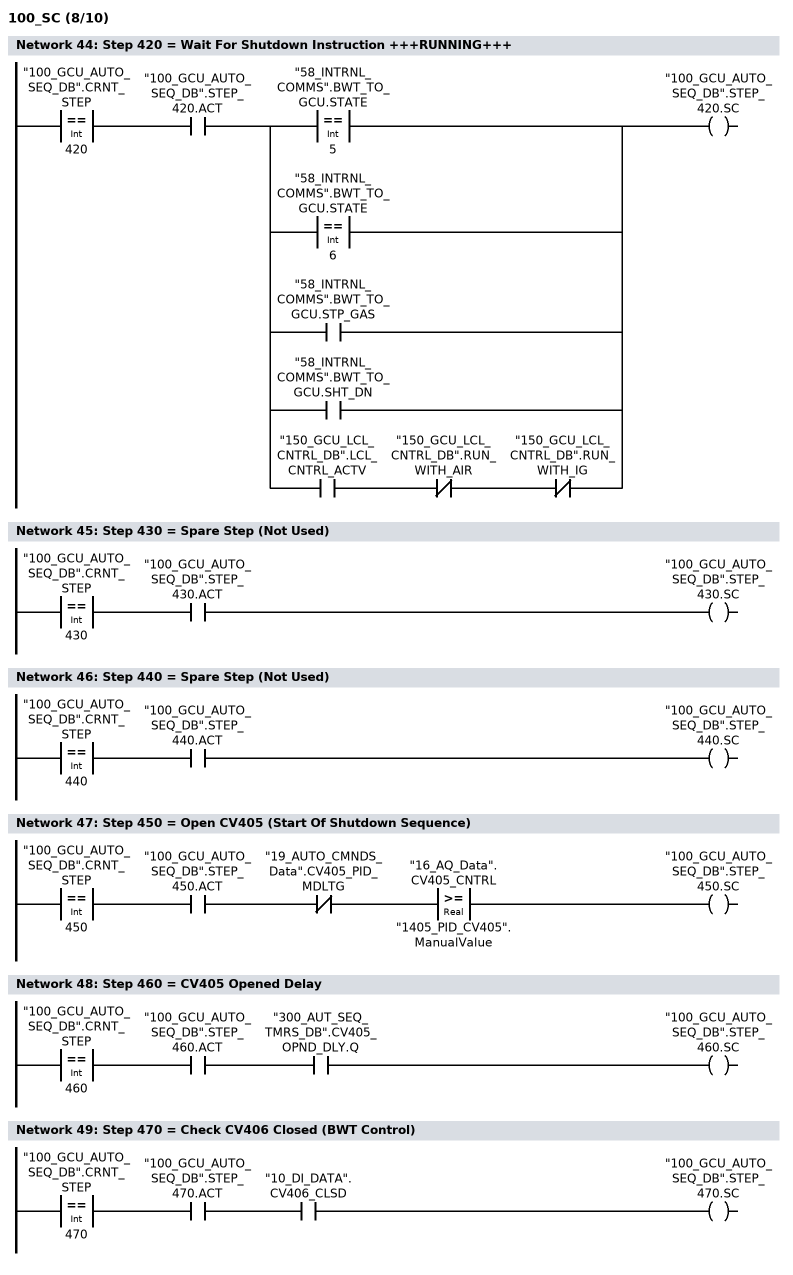
   RUNG wire#powerrail
      { S7_Templates := "SrcType := Int" } EQ_Contact(in1 := "100_GCU_AUTO_SEQ_DB".CRNT_STEP, in2 := 420)
      Contact( "100_GCU_AUTO_SEQ_DB".STEP_420.ACT )
      wire#w1
      { S7_Templates := "SrcType := Int" } EQ_Contact(in1 := "58_INTRNL_COMMS".BWT_TO_GCU.STATE, in2 := 5)
      wire#w2
      Coil( "100_GCU_AUTO_SEQ_DB".STEP_420.SC )
   END_RUNG
   RUNG wire#w1
      { S7_Templates := "SrcType := Int" } EQ_Contact(in1 := "58_INTRNL_COMMS".BWT_TO_GCU.STATE, in2 := 6)
   END_RUNG wire#w2
   RUNG wire#w1
      Contact( "58_INTRNL_COMMS".BWT_TO_GCU.STP_GAS )
   END_RUNG wire#w2
   RUNG wire#w1
      Contact( "58_INTRNL_COMMS".BWT_TO_GCU.SHT_DN )
   END_RUNG wire#w2
   RUNG wire#w1
      Contact( "150_GCU_LCL_CNTRL_DB".LCL_CNTRL_ACTV )
      I_Contact( "150_GCU_LCL_CNTRL_DB".RUN_WITH_AIR )
      I_Contact( "150_GCU_LCL_CNTRL_DB".RUN_WITH_IG )
   END_RUNG wire#w2
   // the same network as SCL:
   "100_GCU_AUTO_SEQ_DB".STEP_420.SC := ("100_GCU_AUTO_SEQ_DB".CRNT_STEP = 420) AND "100_GCU_AUTO_SEQ_DB".STEP_420.ACT AND (("58_INTRNL_COMMS".BWT_TO_GCU.STATE = 5) OR ("58_INTRNL_COMMS".BWT_TO_GCU.STATE = 6) OR "58_INTRNL_COMMS".BWT_TO_GCU.STP_GAS OR "58_INTRNL_COMMS".BWT_TO_GCU.SHT_DN OR ("150_GCU_LCL_CNTRL_DB".LCL_CNTRL_ACTV AND NOT "150_GCU_LCL_CNTRL_DB".RUN_WITH_AIR AND NOT "150_GCU_LCL_CNTRL_DB".RUN_WITH_IG));
END_REGION

REGION Network 45: Step 430 = Spare Step (Not Used)
   RUNG wire#powerrail
      { S7_Templates := "SrcType := Int" } EQ_Contact(in1 := "100_GCU_AUTO_SEQ_DB".CRNT_STEP, in2 := 430)
      Contact( "100_GCU_AUTO_SEQ_DB".STEP_430.ACT )
      Coil( "100_GCU_AUTO_SEQ_DB".STEP_430.SC )
   END_RUNG
   // the same network as SCL:
   "100_GCU_AUTO_SEQ_DB".STEP_430.SC := ("100_GCU_AUTO_SEQ_DB".CRNT_STEP = 430) AND "100_GCU_AUTO_SEQ_DB".STEP_430.ACT;
END_REGION

REGION Network 46: Step 440 = Spare Step (Not Used)
   RUNG wire#powerrail
      { S7_Templates := "SrcType := Int" } EQ_Contact(in1 := "100_GCU_AUTO_SEQ_DB".CRNT_STEP, in2 := 440)
      Contact( "100_GCU_AUTO_SEQ_DB".STEP_440.ACT )
      Coil( "100_GCU_AUTO_SEQ_DB".STEP_440.SC )
   END_RUNG
   // the same network as SCL:
   "100_GCU_AUTO_SEQ_DB".STEP_440.SC := ("100_GCU_AUTO_SEQ_DB".CRNT_STEP = 440) AND "100_GCU_AUTO_SEQ_DB".STEP_440.ACT;
END_REGION

REGION Network 47: Step 450 = Open CV405 (Start Of Shutdown Sequence)
   RUNG wire#powerrail
      { S7_Templates := "SrcType := Int" } EQ_Contact(in1 := "100_GCU_AUTO_SEQ_DB".CRNT_STEP, in2 := 450)
      Contact( "100_GCU_AUTO_SEQ_DB".STEP_450.ACT )
      I_Contact( "19_AUTO_CMNDS_Data".CV405_PID_MDLTG )
      { S7_Templates := "SrcType := Real" } GE_Contact(in1 := "16_AQ_Data".CV405_CNTRL, in2 := "1405_PID_CV405".ManualValue)
      Coil( "100_GCU_AUTO_SEQ_DB".STEP_450.SC )
   END_RUNG
   // the same network as SCL:
   "100_GCU_AUTO_SEQ_DB".STEP_450.SC := ("100_GCU_AUTO_SEQ_DB".CRNT_STEP = 450) AND "100_GCU_AUTO_SEQ_DB".STEP_450.ACT AND NOT "19_AUTO_CMNDS_Data".CV405_PID_MDLTG AND ("16_AQ_Data".CV405_CNTRL >= "1405_PID_CV405".ManualValue);
END_REGION

REGION Network 48: Step 460 = CV405 Opened Delay
   RUNG wire#powerrail
      { S7_Templates := "SrcType := Int" } EQ_Contact(in1 := "100_GCU_AUTO_SEQ_DB".CRNT_STEP, in2 := 460)
      Contact( "100_GCU_AUTO_SEQ_DB".STEP_460.ACT )
      Contact( "300_AUT_SEQ_TMRS_DB".CV405_OPND_DLY.Q )
      Coil( "100_GCU_AUTO_SEQ_DB".STEP_460.SC )
   END_RUNG
   // the same network as SCL:
   "100_GCU_AUTO_SEQ_DB".STEP_460.SC := ("100_GCU_AUTO_SEQ_DB".CRNT_STEP = 460) AND "100_GCU_AUTO_SEQ_DB".STEP_460.ACT AND "300_AUT_SEQ_TMRS_DB".CV405_OPND_DLY.Q;
END_REGION

REGION Network 49: Step 470 = Check CV406 Closed (BWT Control)
   RUNG wire#powerrail
      { S7_Templates := "SrcType := Int" } EQ_Contact(in1 := "100_GCU_AUTO_SEQ_DB".CRNT_STEP, in2 := 470)
      Contact( "100_GCU_AUTO_SEQ_DB".STEP_470.ACT )
      Contact( "10_DI_DATA".CV406_CLSD )
      Coil( "100_GCU_AUTO_SEQ_DB".STEP_470.SC )
   END_RUNG
   // the same network as SCL:
   "100_GCU_AUTO_SEQ_DB".STEP_470.SC := ("100_GCU_AUTO_SEQ_DB".CRNT_STEP = 470) AND "100_GCU_AUTO_SEQ_DB".STEP_470.ACT AND "10_DI_DATA".CV406_CLSD;
END_REGION

REGION Network 50: Step 480 = CV406 Closed Delay & PGC Flush Delay
   // Condition added to whait PGC flush sequence
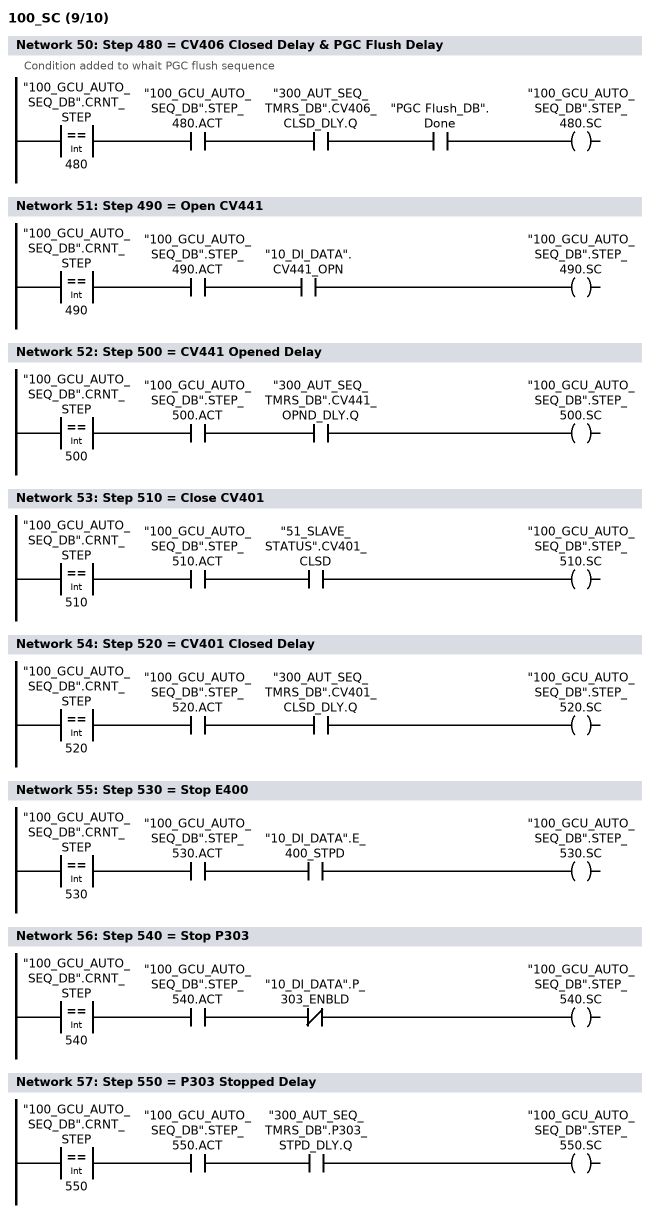
   RUNG wire#powerrail
      { S7_Templates := "SrcType := Int" } EQ_Contact(in1 := "100_GCU_AUTO_SEQ_DB".CRNT_STEP, in2 := 480)
      Contact( "100_GCU_AUTO_SEQ_DB".STEP_480.ACT )
      Contact( "300_AUT_SEQ_TMRS_DB".CV406_CLSD_DLY.Q )
      Contact( "PGC Flush_DB".Done )
      Coil( "100_GCU_AUTO_SEQ_DB".STEP_480.SC )
   END_RUNG
   // the same network as SCL:
   "100_GCU_AUTO_SEQ_DB".STEP_480.SC := ("100_GCU_AUTO_SEQ_DB".CRNT_STEP = 480) AND "100_GCU_AUTO_SEQ_DB".STEP_480.ACT AND "300_AUT_SEQ_TMRS_DB".CV406_CLSD_DLY.Q AND "PGC Flush_DB".Done;
END_REGION

REGION Network 51: Step 490 = Open CV441
   RUNG wire#powerrail
      { S7_Templates := "SrcType := Int" } EQ_Contact(in1 := "100_GCU_AUTO_SEQ_DB".CRNT_STEP, in2 := 490)
      Contact( "100_GCU_AUTO_SEQ_DB".STEP_490.ACT )
      Contact( "10_DI_DATA".CV441_OPN )
      Coil( "100_GCU_AUTO_SEQ_DB".STEP_490.SC )
   END_RUNG
   // the same network as SCL:
   "100_GCU_AUTO_SEQ_DB".STEP_490.SC := ("100_GCU_AUTO_SEQ_DB".CRNT_STEP = 490) AND "100_GCU_AUTO_SEQ_DB".STEP_490.ACT AND "10_DI_DATA".CV441_OPN;
END_REGION

REGION Network 52: Step 500 = CV441 Opened Delay
   RUNG wire#powerrail
      { S7_Templates := "SrcType := Int" } EQ_Contact(in1 := "100_GCU_AUTO_SEQ_DB".CRNT_STEP, in2 := 500)
      Contact( "100_GCU_AUTO_SEQ_DB".STEP_500.ACT )
      Contact( "300_AUT_SEQ_TMRS_DB".CV441_OPND_DLY.Q )
      Coil( "100_GCU_AUTO_SEQ_DB".STEP_500.SC )
   END_RUNG
   // the same network as SCL:
   "100_GCU_AUTO_SEQ_DB".STEP_500.SC := ("100_GCU_AUTO_SEQ_DB".CRNT_STEP = 500) AND "100_GCU_AUTO_SEQ_DB".STEP_500.ACT AND "300_AUT_SEQ_TMRS_DB".CV441_OPND_DLY.Q;
END_REGION

REGION Network 53: Step 510 = Close CV401
   RUNG wire#powerrail
      { S7_Templates := "SrcType := Int" } EQ_Contact(in1 := "100_GCU_AUTO_SEQ_DB".CRNT_STEP, in2 := 510)
      Contact( "100_GCU_AUTO_SEQ_DB".STEP_510.ACT )
      Contact( "51_SLAVE_STATUS".CV401_CLSD )
      Coil( "100_GCU_AUTO_SEQ_DB".STEP_510.SC )
   END_RUNG
   // the same network as SCL:
   "100_GCU_AUTO_SEQ_DB".STEP_510.SC := ("100_GCU_AUTO_SEQ_DB".CRNT_STEP = 510) AND "100_GCU_AUTO_SEQ_DB".STEP_510.ACT AND "51_SLAVE_STATUS".CV401_CLSD;
END_REGION

REGION Network 54: Step 520 = CV401 Closed Delay
   RUNG wire#powerrail
      { S7_Templates := "SrcType := Int" } EQ_Contact(in1 := "100_GCU_AUTO_SEQ_DB".CRNT_STEP, in2 := 520)
      Contact( "100_GCU_AUTO_SEQ_DB".STEP_520.ACT )
      Contact( "300_AUT_SEQ_TMRS_DB".CV401_CLSD_DLY.Q )
      Coil( "100_GCU_AUTO_SEQ_DB".STEP_520.SC )
   END_RUNG
   // the same network as SCL:
   "100_GCU_AUTO_SEQ_DB".STEP_520.SC := ("100_GCU_AUTO_SEQ_DB".CRNT_STEP = 520) AND "100_GCU_AUTO_SEQ_DB".STEP_520.ACT AND "300_AUT_SEQ_TMRS_DB".CV401_CLSD_DLY.Q;
END_REGION

REGION Network 55: Step 530 = Stop E400
   RUNG wire#powerrail
      { S7_Templates := "SrcType := Int" } EQ_Contact(in1 := "100_GCU_AUTO_SEQ_DB".CRNT_STEP, in2 := 530)
      Contact( "100_GCU_AUTO_SEQ_DB".STEP_530.ACT )
      Contact( "10_DI_DATA".E_400_STPD )
      Coil( "100_GCU_AUTO_SEQ_DB".STEP_530.SC )
   END_RUNG
   // the same network as SCL:
   "100_GCU_AUTO_SEQ_DB".STEP_530.SC := ("100_GCU_AUTO_SEQ_DB".CRNT_STEP = 530) AND "100_GCU_AUTO_SEQ_DB".STEP_530.ACT AND "10_DI_DATA".E_400_STPD;
END_REGION

REGION Network 56: Step 540 = Stop P303
   RUNG wire#powerrail
      { S7_Templates := "SrcType := Int" } EQ_Contact(in1 := "100_GCU_AUTO_SEQ_DB".CRNT_STEP, in2 := 540)
      Contact( "100_GCU_AUTO_SEQ_DB".STEP_540.ACT )
      I_Contact( "10_DI_DATA".P_303_ENBLD )
      Coil( "100_GCU_AUTO_SEQ_DB".STEP_540.SC )
   END_RUNG
   // the same network as SCL:
   "100_GCU_AUTO_SEQ_DB".STEP_540.SC := ("100_GCU_AUTO_SEQ_DB".CRNT_STEP = 540) AND "100_GCU_AUTO_SEQ_DB".STEP_540.ACT AND NOT "10_DI_DATA".P_303_ENBLD;
END_REGION

REGION Network 57: Step 550 = P303 Stopped Delay
   RUNG wire#powerrail
      { S7_Templates := "SrcType := Int" } EQ_Contact(in1 := "100_GCU_AUTO_SEQ_DB".CRNT_STEP, in2 := 550)
      Contact( "100_GCU_AUTO_SEQ_DB".STEP_550.ACT )
      Contact( "300_AUT_SEQ_TMRS_DB".P303_STPD_DLY.Q )
      Coil( "100_GCU_AUTO_SEQ_DB".STEP_550.SC )
   END_RUNG
   // the same network as SCL:
   "100_GCU_AUTO_SEQ_DB".STEP_550.SC := ("100_GCU_AUTO_SEQ_DB".CRNT_STEP = 550) AND "100_GCU_AUTO_SEQ_DB".STEP_550.ACT AND "300_AUT_SEQ_TMRS_DB".P303_STPD_DLY.Q;
END_REGION

REGION Network 58: Step 560 = Wait For PIT416 <0.01bar
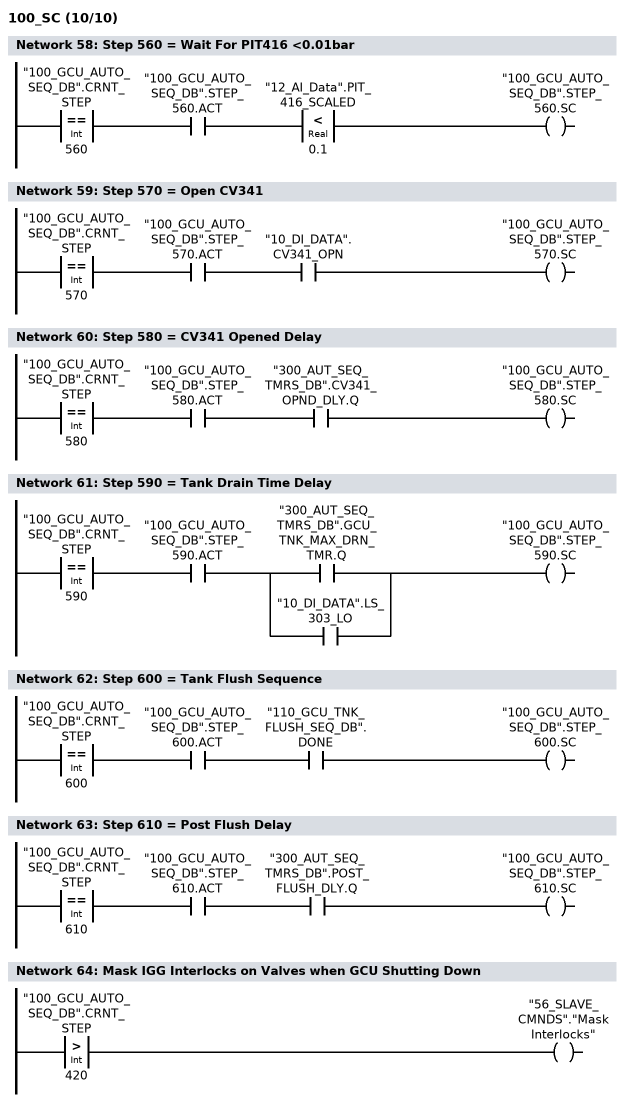
   RUNG wire#powerrail
      { S7_Templates := "SrcType := Int" } EQ_Contact(in1 := "100_GCU_AUTO_SEQ_DB".CRNT_STEP, in2 := 560)
      Contact( "100_GCU_AUTO_SEQ_DB".STEP_560.ACT )
      { S7_Templates := "SrcType := Real" } LT_Contact(in1 := "12_AI_Data".PIT_416_SCALED, in2 := 0.1)
      Coil( "100_GCU_AUTO_SEQ_DB".STEP_560.SC )
   END_RUNG
   // the same network as SCL:
   "100_GCU_AUTO_SEQ_DB".STEP_560.SC := ("100_GCU_AUTO_SEQ_DB".CRNT_STEP = 560) AND "100_GCU_AUTO_SEQ_DB".STEP_560.ACT AND ("12_AI_Data".PIT_416_SCALED < 0.1);
END_REGION

REGION Network 59: Step 570 = Open CV341
   RUNG wire#powerrail
      { S7_Templates := "SrcType := Int" } EQ_Contact(in1 := "100_GCU_AUTO_SEQ_DB".CRNT_STEP, in2 := 570)
      Contact( "100_GCU_AUTO_SEQ_DB".STEP_570.ACT )
      Contact( "10_DI_DATA".CV341_OPN )
      Coil( "100_GCU_AUTO_SEQ_DB".STEP_570.SC )
   END_RUNG
   // the same network as SCL:
   "100_GCU_AUTO_SEQ_DB".STEP_570.SC := ("100_GCU_AUTO_SEQ_DB".CRNT_STEP = 570) AND "100_GCU_AUTO_SEQ_DB".STEP_570.ACT AND "10_DI_DATA".CV341_OPN;
END_REGION

REGION Network 60: Step 580 = CV341 Opened Delay
   RUNG wire#powerrail
      { S7_Templates := "SrcType := Int" } EQ_Contact(in1 := "100_GCU_AUTO_SEQ_DB".CRNT_STEP, in2 := 580)
      Contact( "100_GCU_AUTO_SEQ_DB".STEP_580.ACT )
      Contact( "300_AUT_SEQ_TMRS_DB".CV341_OPND_DLY.Q )
      Coil( "100_GCU_AUTO_SEQ_DB".STEP_580.SC )
   END_RUNG
   // the same network as SCL:
   "100_GCU_AUTO_SEQ_DB".STEP_580.SC := ("100_GCU_AUTO_SEQ_DB".CRNT_STEP = 580) AND "100_GCU_AUTO_SEQ_DB".STEP_580.ACT AND "300_AUT_SEQ_TMRS_DB".CV341_OPND_DLY.Q;
END_REGION

REGION Network 61: Step 590 = Tank Drain Time Delay
   RUNG wire#powerrail
      { S7_Templates := "SrcType := Int" } EQ_Contact(in1 := "100_GCU_AUTO_SEQ_DB".CRNT_STEP, in2 := 590)
      Contact( "100_GCU_AUTO_SEQ_DB".STEP_590.ACT )
      wire#w1
      Contact( "300_AUT_SEQ_TMRS_DB".GCU_TNK_MAX_DRN_TMR.Q )
      wire#w2
      Coil( "100_GCU_AUTO_SEQ_DB".STEP_590.SC )
   END_RUNG
   RUNG wire#w1
      Contact( "10_DI_DATA".LS_303_LO )
   END_RUNG wire#w2
   // the same network as SCL:
   "100_GCU_AUTO_SEQ_DB".STEP_590.SC := ("100_GCU_AUTO_SEQ_DB".CRNT_STEP = 590) AND "100_GCU_AUTO_SEQ_DB".STEP_590.ACT AND ("300_AUT_SEQ_TMRS_DB".GCU_TNK_MAX_DRN_TMR.Q OR "10_DI_DATA".LS_303_LO);
END_REGION

REGION Network 62: Step 600 = Tank Flush Sequence
   RUNG wire#powerrail
      { S7_Templates := "SrcType := Int" } EQ_Contact(in1 := "100_GCU_AUTO_SEQ_DB".CRNT_STEP, in2 := 600)
      Contact( "100_GCU_AUTO_SEQ_DB".STEP_600.ACT )
      Contact( "110_GCU_TNK_FLUSH_SEQ_DB".DONE )
      Coil( "100_GCU_AUTO_SEQ_DB".STEP_600.SC )
   END_RUNG
   // the same network as SCL:
   "100_GCU_AUTO_SEQ_DB".STEP_600.SC := ("100_GCU_AUTO_SEQ_DB".CRNT_STEP = 600) AND "100_GCU_AUTO_SEQ_DB".STEP_600.ACT AND "110_GCU_TNK_FLUSH_SEQ_DB".DONE;
END_REGION

REGION Network 63: Step 610 = Post Flush Delay
   RUNG wire#powerrail
      { S7_Templates := "SrcType := Int" } EQ_Contact(in1 := "100_GCU_AUTO_SEQ_DB".CRNT_STEP, in2 := 610)
      Contact( "100_GCU_AUTO_SEQ_DB".STEP_610.ACT )
      Contact( "300_AUT_SEQ_TMRS_DB".POST_FLUSH_DLY.Q )
      Coil( "100_GCU_AUTO_SEQ_DB".STEP_610.SC )
   END_RUNG
   // the same network as SCL:
   "100_GCU_AUTO_SEQ_DB".STEP_610.SC := ("100_GCU_AUTO_SEQ_DB".CRNT_STEP = 610) AND "100_GCU_AUTO_SEQ_DB".STEP_610.ACT AND "300_AUT_SEQ_TMRS_DB".POST_FLUSH_DLY.Q;
END_REGION

REGION Network 64: Mask IGG Interlocks on Valves when GCU Shutting Down
   RUNG wire#powerrail
      { S7_Templates := "SrcType := Int" } GT_Contact(in1 := "100_GCU_AUTO_SEQ_DB".CRNT_STEP, in2 := 420)
      Coil( "56_SLAVE_CMNDS"."Mask Interlocks" )
   END_RUNG
   // the same network as SCL:
   "56_SLAVE_CMNDS"."Mask Interlocks" := "100_GCU_AUTO_SEQ_DB".CRNT_STEP > 420;
END_REGION
END_FUNCTION

FUNCTION "101_SP_CNFG" : Void   // FC101, LAD
TITLE = Setpoint Configuration
{ S7_Optimized_Access := 'TRUE' }
AUTHOR : JRS
VERSION : 0.1
// For configuring setpoints during automatic operation
   VAR_TEMP   // added for the SCL form of the ladder/FBD networks
      _w1 : Bool;
   END_VAR
BEGIN

REGION Network 1: LIT304
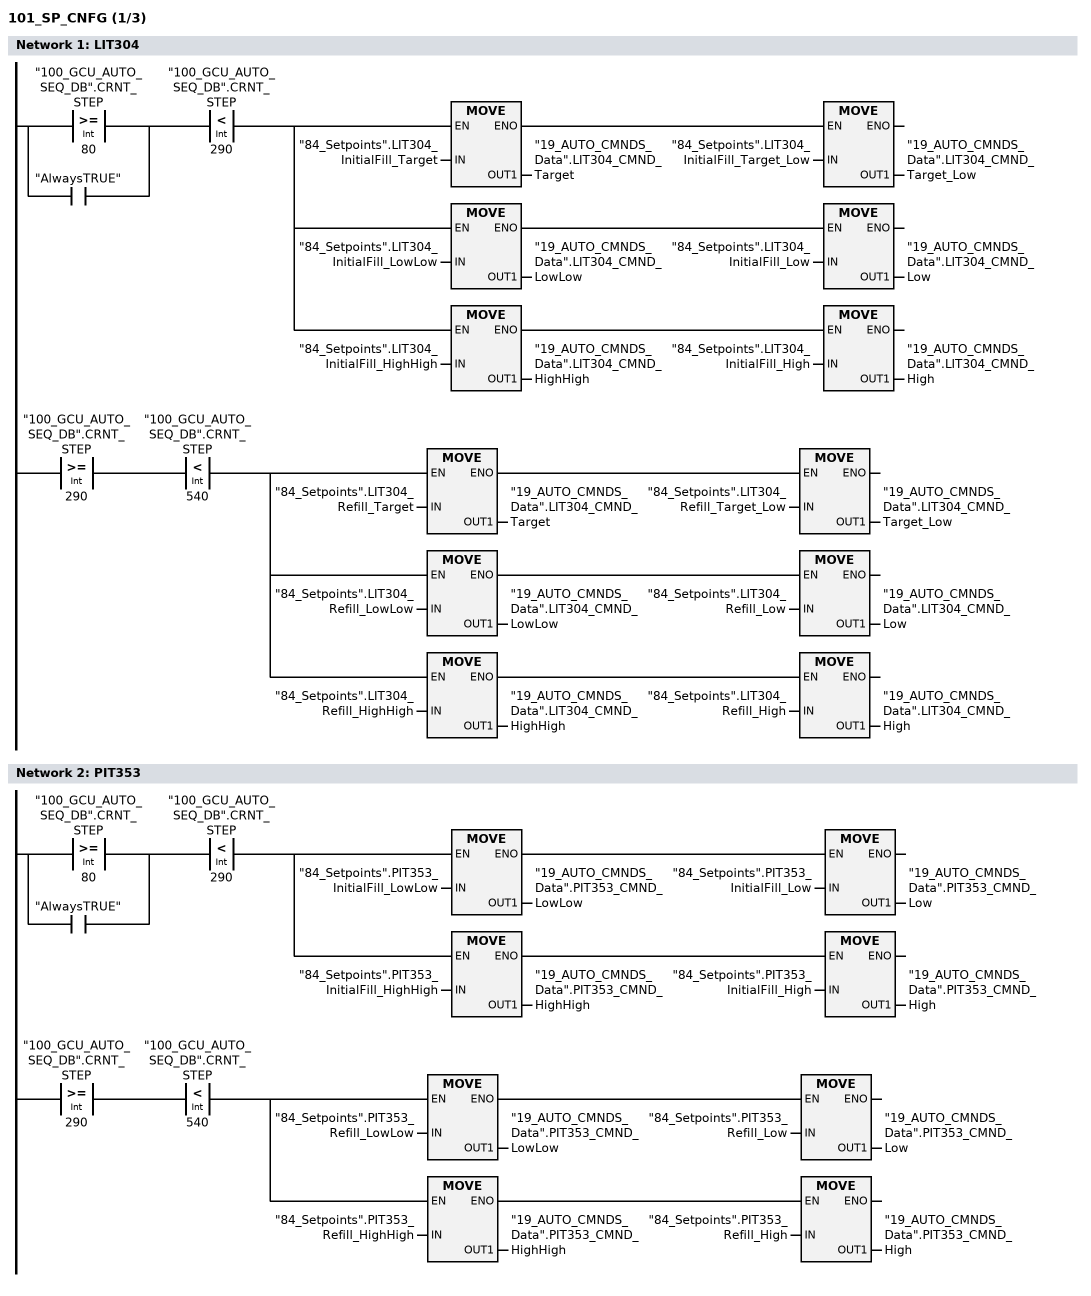
   RUNG wire#powerrail
      { S7_Templates := "SrcType := Int" } GE_Contact(in1 := "100_GCU_AUTO_SEQ_DB".CRNT_STEP, in2 := 80)
      wire#w1
      { S7_Templates := "SrcType := Int" } LT_Contact(in1 := "100_GCU_AUTO_SEQ_DB".CRNT_STEP, in2 := 290)
      wire#w2
      Move(in := "84_Setpoints".LIT304_InitialFill_Target, out1 => "19_AUTO_CMNDS_Data".LIT304_CMND_Target)
      Move(in := "84_Setpoints".LIT304_InitialFill_Target_Low, out1 => "19_AUTO_CMNDS_Data".LIT304_CMND_Target_Low)
   END_RUNG
   RUNG wire#powerrail
      Contact( "AlwaysTRUE" )
   END_RUNG wire#w1
   RUNG wire#w2
      Move(in := "84_Setpoints".LIT304_InitialFill_LowLow, out1 => "19_AUTO_CMNDS_Data".LIT304_CMND_LowLow)
      Move(in := "84_Setpoints".LIT304_InitialFill_Low, out1 => "19_AUTO_CMNDS_Data".LIT304_CMND_Low)
   END_RUNG
   RUNG wire#w2
      Move(in := "84_Setpoints".LIT304_InitialFill_HighHigh, out1 => "19_AUTO_CMNDS_Data".LIT304_CMND_HighHigh)
      Move(in := "84_Setpoints".LIT304_InitialFill_High, out1 => "19_AUTO_CMNDS_Data".LIT304_CMND_High)
   END_RUNG
   RUNG wire#powerrail
      { S7_Templates := "SrcType := Int" } GE_Contact(in1 := "100_GCU_AUTO_SEQ_DB".CRNT_STEP, in2 := 290)
      { S7_Templates := "SrcType := Int" } LT_Contact(in1 := "100_GCU_AUTO_SEQ_DB".CRNT_STEP, in2 := 540)
      wire#w3
      Move(in := "84_Setpoints".LIT304_Refill_Target, out1 => "19_AUTO_CMNDS_Data".LIT304_CMND_Target)
      Move(in := "84_Setpoints".LIT304_Refill_Target_Low, out1 => "19_AUTO_CMNDS_Data".LIT304_CMND_Target_Low)
   END_RUNG
   RUNG wire#w3
      Move(in := "84_Setpoints".LIT304_Refill_LowLow, out1 => "19_AUTO_CMNDS_Data".LIT304_CMND_LowLow)
      Move(in := "84_Setpoints".LIT304_Refill_Low, out1 => "19_AUTO_CMNDS_Data".LIT304_CMND_Low)
   END_RUNG
   RUNG wire#w3
      Move(in := "84_Setpoints".LIT304_Refill_HighHigh, out1 => "19_AUTO_CMNDS_Data".LIT304_CMND_HighHigh)
      Move(in := "84_Setpoints".LIT304_Refill_High, out1 => "19_AUTO_CMNDS_Data".LIT304_CMND_High)
   END_RUNG
   // the same network as SCL:
   IF (("100_GCU_AUTO_SEQ_DB".CRNT_STEP >= 80) OR "AlwaysTRUE") AND ("100_GCU_AUTO_SEQ_DB".CRNT_STEP < 290) THEN
       "19_AUTO_CMNDS_Data".LIT304_CMND_Target := "84_Setpoints".LIT304_InitialFill_Target;
       "19_AUTO_CMNDS_Data".LIT304_CMND_Target_Low := "84_Setpoints".LIT304_InitialFill_Target_Low;
       "19_AUTO_CMNDS_Data".LIT304_CMND_LowLow := "84_Setpoints".LIT304_InitialFill_LowLow;
       "19_AUTO_CMNDS_Data".LIT304_CMND_Low := "84_Setpoints".LIT304_InitialFill_Low;
       "19_AUTO_CMNDS_Data".LIT304_CMND_HighHigh := "84_Setpoints".LIT304_InitialFill_HighHigh;
       "19_AUTO_CMNDS_Data".LIT304_CMND_High := "84_Setpoints".LIT304_InitialFill_High;
   END_IF;
   IF ("100_GCU_AUTO_SEQ_DB".CRNT_STEP >= 290) AND ("100_GCU_AUTO_SEQ_DB".CRNT_STEP < 540) THEN
       "19_AUTO_CMNDS_Data".LIT304_CMND_Target := "84_Setpoints".LIT304_Refill_Target;
       "19_AUTO_CMNDS_Data".LIT304_CMND_Target_Low := "84_Setpoints".LIT304_Refill_Target_Low;
       "19_AUTO_CMNDS_Data".LIT304_CMND_LowLow := "84_Setpoints".LIT304_Refill_LowLow;
       "19_AUTO_CMNDS_Data".LIT304_CMND_Low := "84_Setpoints".LIT304_Refill_Low;
       "19_AUTO_CMNDS_Data".LIT304_CMND_HighHigh := "84_Setpoints".LIT304_Refill_HighHigh;
       "19_AUTO_CMNDS_Data".LIT304_CMND_High := "84_Setpoints".LIT304_Refill_High;
   END_IF;
END_REGION

REGION Network 2: PIT353
   RUNG wire#powerrail
      { S7_Templates := "SrcType := Int" } GE_Contact(in1 := "100_GCU_AUTO_SEQ_DB".CRNT_STEP, in2 := 80)
      wire#w1
      { S7_Templates := "SrcType := Int" } LT_Contact(in1 := "100_GCU_AUTO_SEQ_DB".CRNT_STEP, in2 := 290)
      wire#w2
      Move(in := "84_Setpoints".PIT353_InitialFill_LowLow, out1 => "19_AUTO_CMNDS_Data".PIT353_CMND_LowLow)
      Move(in := "84_Setpoints".PIT353_InitialFill_Low, out1 => "19_AUTO_CMNDS_Data".PIT353_CMND_Low)
   END_RUNG
   RUNG wire#powerrail
      Contact( "AlwaysTRUE" )
   END_RUNG wire#w1
   RUNG wire#w2
      Move(in := "84_Setpoints".PIT353_InitialFill_HighHigh, out1 => "19_AUTO_CMNDS_Data".PIT353_CMND_HighHigh)
      Move(in := "84_Setpoints".PIT353_InitialFill_High, out1 => "19_AUTO_CMNDS_Data".PIT353_CMND_High)
   END_RUNG
   RUNG wire#powerrail
      { S7_Templates := "SrcType := Int" } GE_Contact(in1 := "100_GCU_AUTO_SEQ_DB".CRNT_STEP, in2 := 290)
      { S7_Templates := "SrcType := Int" } LT_Contact(in1 := "100_GCU_AUTO_SEQ_DB".CRNT_STEP, in2 := 540)
      wire#w3
      Move(in := "84_Setpoints".PIT353_Refill_LowLow, out1 => "19_AUTO_CMNDS_Data".PIT353_CMND_LowLow)
      Move(in := "84_Setpoints".PIT353_Refill_Low, out1 => "19_AUTO_CMNDS_Data".PIT353_CMND_Low)
   END_RUNG
   RUNG wire#w3
      Move(in := "84_Setpoints".PIT353_Refill_HighHigh, out1 => "19_AUTO_CMNDS_Data".PIT353_CMND_HighHigh)
      Move(in := "84_Setpoints".PIT353_Refill_High, out1 => "19_AUTO_CMNDS_Data".PIT353_CMND_High)
   END_RUNG
   // the same network as SCL:
   IF (("100_GCU_AUTO_SEQ_DB".CRNT_STEP >= 80) OR "AlwaysTRUE") AND ("100_GCU_AUTO_SEQ_DB".CRNT_STEP < 290) THEN
       "19_AUTO_CMNDS_Data".PIT353_CMND_LowLow := "84_Setpoints".PIT353_InitialFill_LowLow;
       "19_AUTO_CMNDS_Data".PIT353_CMND_Low := "84_Setpoints".PIT353_InitialFill_Low;
       "19_AUTO_CMNDS_Data".PIT353_CMND_HighHigh := "84_Setpoints".PIT353_InitialFill_HighHigh;
       "19_AUTO_CMNDS_Data".PIT353_CMND_High := "84_Setpoints".PIT353_InitialFill_High;
   END_IF;
   IF ("100_GCU_AUTO_SEQ_DB".CRNT_STEP >= 290) AND ("100_GCU_AUTO_SEQ_DB".CRNT_STEP < 540) THEN
       "19_AUTO_CMNDS_Data".PIT353_CMND_LowLow := "84_Setpoints".PIT353_Refill_LowLow;
       "19_AUTO_CMNDS_Data".PIT353_CMND_Low := "84_Setpoints".PIT353_Refill_Low;
       "19_AUTO_CMNDS_Data".PIT353_CMND_HighHigh := "84_Setpoints".PIT353_Refill_HighHigh;
       "19_AUTO_CMNDS_Data".PIT353_CMND_High := "84_Setpoints".PIT353_Refill_High;
   END_IF;
END_REGION

REGION Network 3: PIT358
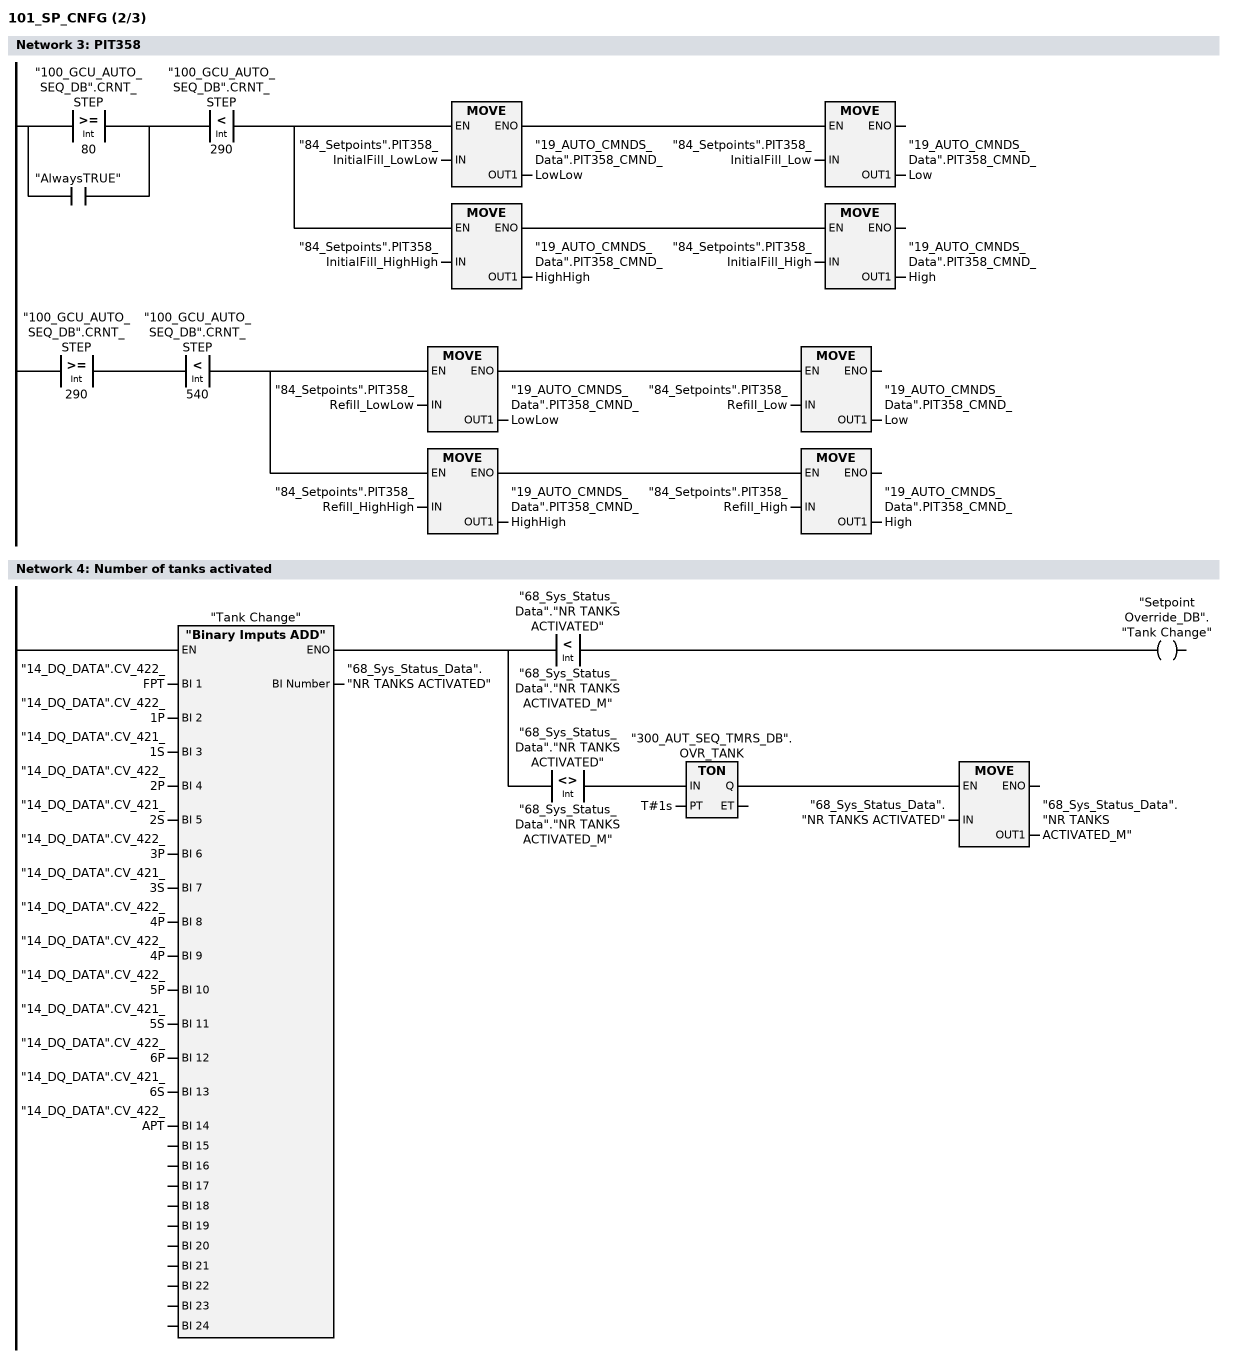
   RUNG wire#powerrail
      { S7_Templates := "SrcType := Int" } GE_Contact(in1 := "100_GCU_AUTO_SEQ_DB".CRNT_STEP, in2 := 80)
      wire#w1
      { S7_Templates := "SrcType := Int" } LT_Contact(in1 := "100_GCU_AUTO_SEQ_DB".CRNT_STEP, in2 := 290)
      wire#w2
      Move(in := "84_Setpoints".PIT358_InitialFill_LowLow, out1 => "19_AUTO_CMNDS_Data".PIT358_CMND_LowLow)
      Move(in := "84_Setpoints".PIT358_InitialFill_Low, out1 => "19_AUTO_CMNDS_Data".PIT358_CMND_Low)
   END_RUNG
   RUNG wire#powerrail
      Contact( "AlwaysTRUE" )
   END_RUNG wire#w1
   RUNG wire#w2
      Move(in := "84_Setpoints".PIT358_InitialFill_HighHigh, out1 => "19_AUTO_CMNDS_Data".PIT358_CMND_HighHigh)
      Move(in := "84_Setpoints".PIT358_InitialFill_High, out1 => "19_AUTO_CMNDS_Data".PIT358_CMND_High)
   END_RUNG
   RUNG wire#powerrail
      { S7_Templates := "SrcType := Int" } GE_Contact(in1 := "100_GCU_AUTO_SEQ_DB".CRNT_STEP, in2 := 290)
      { S7_Templates := "SrcType := Int" } LT_Contact(in1 := "100_GCU_AUTO_SEQ_DB".CRNT_STEP, in2 := 540)
      wire#w3
      Move(in := "84_Setpoints".PIT358_Refill_LowLow, out1 => "19_AUTO_CMNDS_Data".PIT358_CMND_LowLow)
      Move(in := "84_Setpoints".PIT358_Refill_Low, out1 => "19_AUTO_CMNDS_Data".PIT358_CMND_Low)
   END_RUNG
   RUNG wire#w3
      Move(in := "84_Setpoints".PIT358_Refill_HighHigh, out1 => "19_AUTO_CMNDS_Data".PIT358_CMND_HighHigh)
      Move(in := "84_Setpoints".PIT358_Refill_High, out1 => "19_AUTO_CMNDS_Data".PIT358_CMND_High)
   END_RUNG
   // the same network as SCL:
   IF (("100_GCU_AUTO_SEQ_DB".CRNT_STEP >= 80) OR "AlwaysTRUE") AND ("100_GCU_AUTO_SEQ_DB".CRNT_STEP < 290) THEN
       "19_AUTO_CMNDS_Data".PIT358_CMND_LowLow := "84_Setpoints".PIT358_InitialFill_LowLow;
       "19_AUTO_CMNDS_Data".PIT358_CMND_Low := "84_Setpoints".PIT358_InitialFill_Low;
       "19_AUTO_CMNDS_Data".PIT358_CMND_HighHigh := "84_Setpoints".PIT358_InitialFill_HighHigh;
       "19_AUTO_CMNDS_Data".PIT358_CMND_High := "84_Setpoints".PIT358_InitialFill_High;
   END_IF;
   IF ("100_GCU_AUTO_SEQ_DB".CRNT_STEP >= 290) AND ("100_GCU_AUTO_SEQ_DB".CRNT_STEP < 540) THEN
       "19_AUTO_CMNDS_Data".PIT358_CMND_LowLow := "84_Setpoints".PIT358_Refill_LowLow;
       "19_AUTO_CMNDS_Data".PIT358_CMND_Low := "84_Setpoints".PIT358_Refill_Low;
       "19_AUTO_CMNDS_Data".PIT358_CMND_HighHigh := "84_Setpoints".PIT358_Refill_HighHigh;
       "19_AUTO_CMNDS_Data".PIT358_CMND_High := "84_Setpoints".PIT358_Refill_High;
   END_IF;
END_REGION

REGION Network 4: Number of tanks activated
   "Tank Change"("BI 1" := "14_DQ_DATA".CV_422_FPT,   // "Binary Imputs ADD"
                 "BI 2" := "14_DQ_DATA".CV_422_1P,
                 "BI 3" := "14_DQ_DATA".CV_421_1S,
                 "BI 4" := "14_DQ_DATA".CV_422_2P,
                 "BI 5" := "14_DQ_DATA".CV_421_2S,
                 "BI 6" := "14_DQ_DATA".CV_422_3P,
                 "BI 7" := "14_DQ_DATA".CV_421_3S,
                 "BI 8" := "14_DQ_DATA".CV_422_4P,
                 "BI 9" := "14_DQ_DATA".CV_422_4P,
                 "BI 10" := "14_DQ_DATA".CV_422_5P,
                 "BI 11" := "14_DQ_DATA".CV_421_5S,
                 "BI 12" := "14_DQ_DATA".CV_422_6P,
                 "BI 13" := "14_DQ_DATA".CV_421_6S,
                 "BI 14" := "14_DQ_DATA".CV_422_APT,
                 "BI Number" => "68_Sys_Status_Data"."NR TANKS ACTIVATED",
                 ENO => #_w1);
   "Setpoint Override_DB"."Tank Change" := #_w1 AND ("68_Sys_Status_Data"."NR TANKS ACTIVATED" < "68_Sys_Status_Data"."NR TANKS ACTIVATED_M");
   "300_AUT_SEQ_TMRS_DB".OVR_TANK.TON(IN := #_w1 AND ("68_Sys_Status_Data"."NR TANKS ACTIVATED" <> "68_Sys_Status_Data"."NR TANKS ACTIVATED_M"),
                           PT := T#1s);
   IF "300_AUT_SEQ_TMRS_DB".OVR_TANK.Q THEN
       "68_Sys_Status_Data"."NR TANKS ACTIVATED_M" := "68_Sys_Status_Data"."NR TANKS ACTIVATED";
   END_IF;
END_REGION

REGION Network 5: Pressure target override to safe conditions
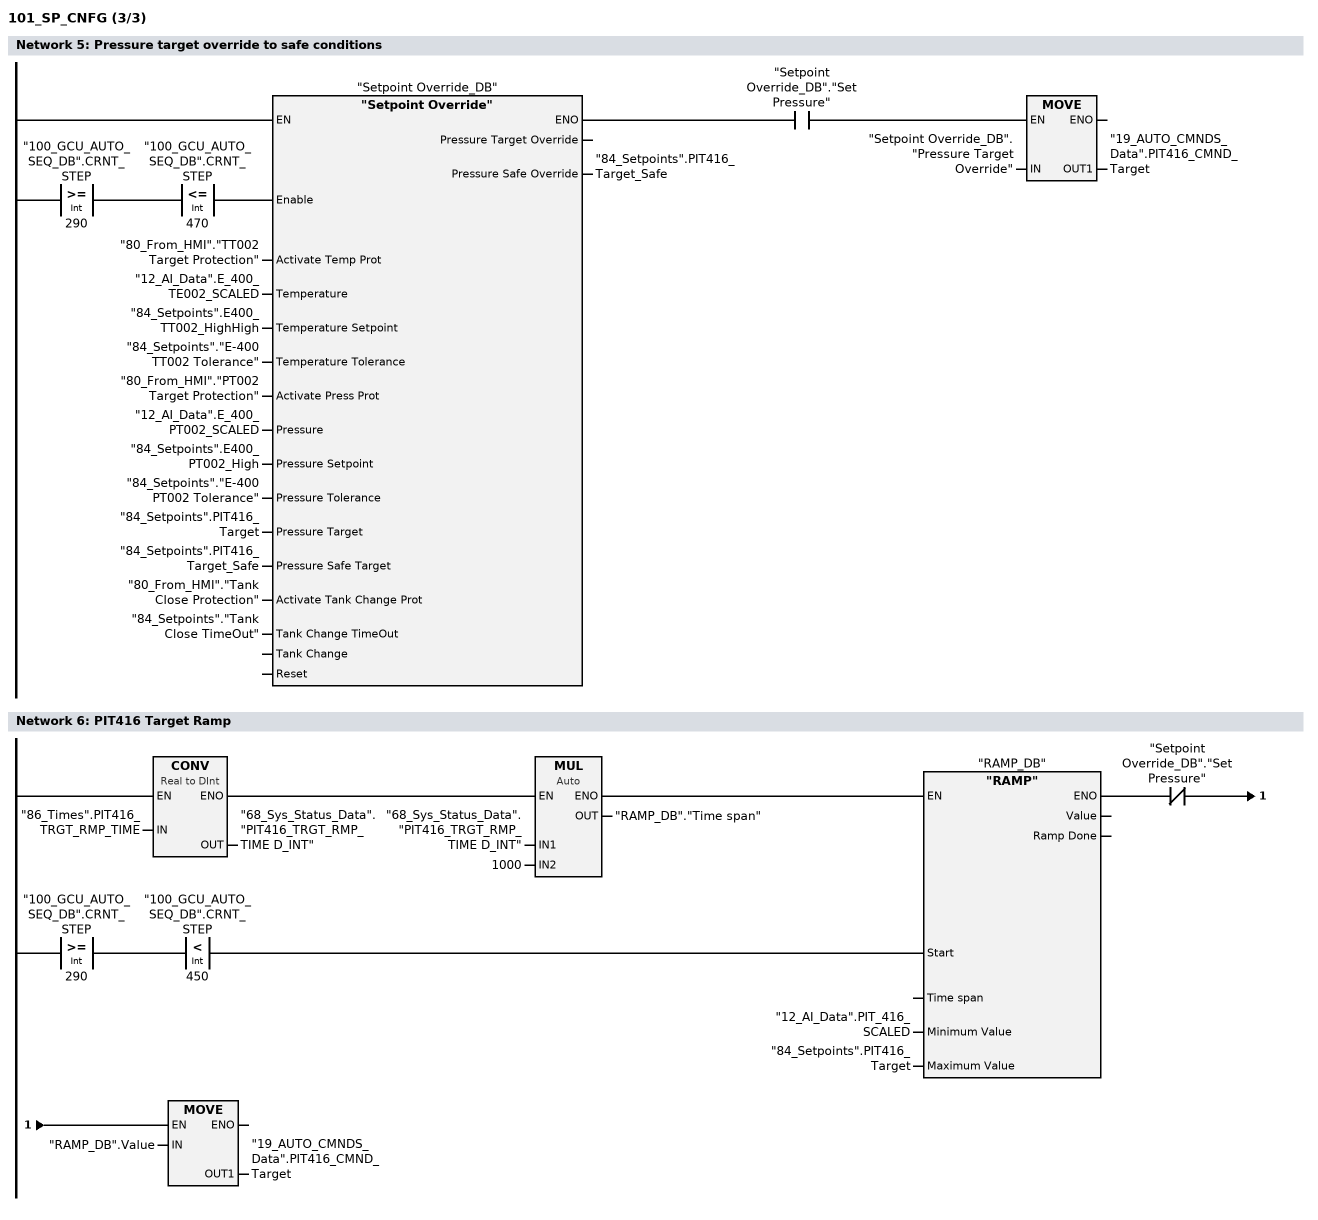
   RUNG wire#powerrail
      "Setpoint Override_DB"(Enable := wire#w1, "Activate Temp Prot" := "80_From_HMI"."TT002 Target Protection", Temperature := "12_AI_Data".E_400_TE002_SCALED, "Temperature Setpoint" := "84_Setpoints".E400_TT002_HighHigh, "Temperature Tolerance" := "84_Setpoints"."E-400 TT002 Tolerance", "Activate Press Prot" := "80_From_HMI"."PT002 Target Protection", Pressure := "12_AI_Data".E_400_PT002_SCALED, "Pressure Setpoint" := "84_Setpoints".E400_PT002_High, "Pressure Tolerance" := "84_Setpoints"."E-400 PT002 Tolerance", "Pressure Target" := "84_Setpoints".PIT416_Target, "Pressure Safe Target" := "84_Setpoints".PIT416_Target_Safe, "Activate Tank Change Prot" := "80_From_HMI"."Tank Close Protection", "Tank Change TimeOut" := "84_Setpoints"."Tank Close TimeOut", "Tank Change" :=, Reset :=, "Pressure Target Override" =>, "Pressure Safe Override" => "84_Setpoints".PIT416_Target_Safe)
      Contact( "Setpoint Override_DB"."Set Pressure" )
      Move(in := "Setpoint Override_DB"."Pressure Target Override", out1 => "19_AUTO_CMNDS_Data".PIT416_CMND_Target)
   END_RUNG
   RUNG wire#powerrail
      { S7_Templates := "SrcType := Int" } GE_Contact(in1 := "100_GCU_AUTO_SEQ_DB".CRNT_STEP, in2 := 290)